REGION Network 26: Check Values
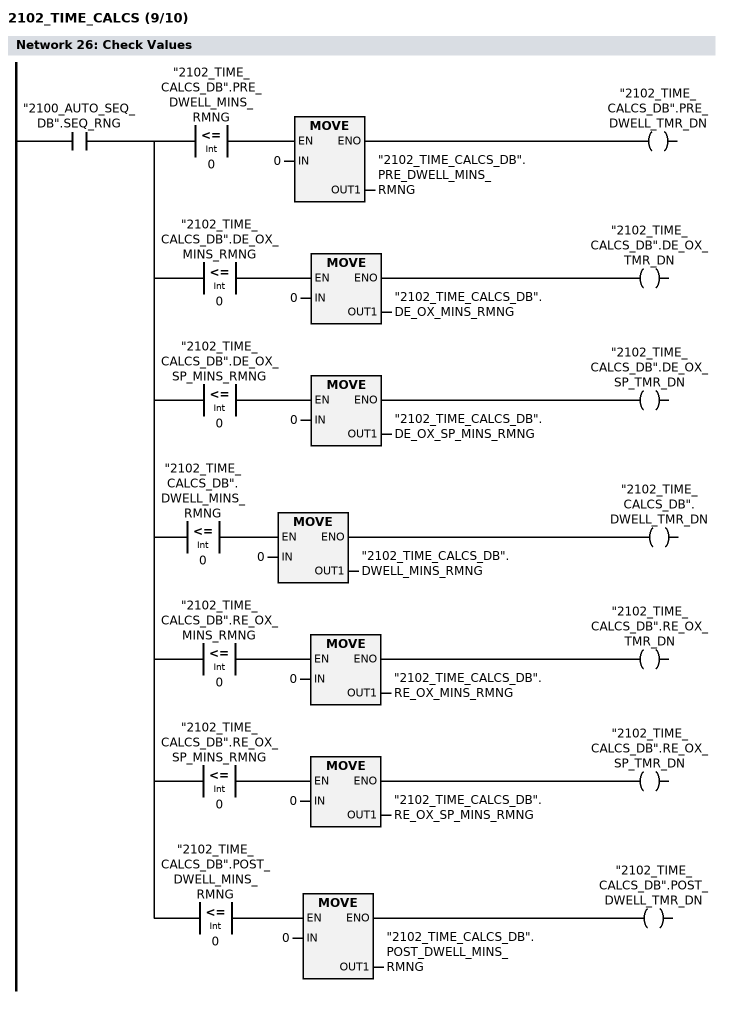
   RUNG wire#powerrail
      Contact( "2100_AUTO_SEQ_DB".SEQ_RNG )
      wire#w1
      { S7_Templates := "SrcType := Int" } LE_Contact(in1 := "2102_TIME_CALCS_DB".PRE_DWELL_MINS_RMNG, in2 := 0)
      Move(in := 0, out1 => "2102_TIME_CALCS_DB".PRE_DWELL_MINS_RMNG)
      Coil( "2102_TIME_CALCS_DB".PRE_DWELL_TMR_DN )
   END_RUNG
   RUNG wire#w1
      { S7_Templates := "SrcType := Int" } LE_Contact(in1 := "2102_TIME_CALCS_DB".DE_OX_MINS_RMNG, in2 := 0)
      Move(in := 0, out1 => "2102_TIME_CALCS_DB".DE_OX_MINS_RMNG)
      Coil( "2102_TIME_CALCS_DB".DE_OX_TMR_DN )
   END_RUNG
   RUNG wire#w1
      { S7_Templates := "SrcType := Int" } LE_Contact(in1 := "2102_TIME_CALCS_DB".DE_OX_SP_MINS_RMNG, in2 := 0)
      Move(in := 0, out1 => "2102_TIME_CALCS_DB".DE_OX_SP_MINS_RMNG)
      Coil( "2102_TIME_CALCS_DB".DE_OX_SP_TMR_DN )
   END_RUNG
   RUNG wire#w1
      { S7_Templates := "SrcType := Int" } LE_Contact(in1 := "2102_TIME_CALCS_DB".DWELL_MINS_RMNG, in2 := 0)
      Move(in := 0, out1 => "2102_TIME_CALCS_DB".DWELL_MINS_RMNG)
      Coil( "2102_TIME_CALCS_DB".DWELL_TMR_DN )
   END_RUNG
   RUNG wire#w1
      { S7_Templates := "SrcType := Int" } LE_Contact(in1 := "2102_TIME_CALCS_DB".RE_OX_MINS_RMNG, in2 := 0)
      Move(in := 0, out1 => "2102_TIME_CALCS_DB".RE_OX_MINS_RMNG)
      Coil( "2102_TIME_CALCS_DB".RE_OX_TMR_DN )
   END_RUNG
   RUNG wire#w1
      { S7_Templates := "SrcType := Int" } LE_Contact(in1 := "2102_TIME_CALCS_DB".RE_OX_SP_MINS_RMNG, in2 := 0)
      Move(in := 0, out1 => "2102_TIME_CALCS_DB".RE_OX_SP_MINS_RMNG)
      Coil( "2102_TIME_CALCS_DB".RE_OX_SP_TMR_DN )
   END_RUNG
   RUNG wire#w1
      { S7_Templates := "SrcType := Int" } LE_Contact(in1 := "2102_TIME_CALCS_DB".POST_DWELL_MINS_RMNG, in2 := 0)
      Move(in := 0, out1 => "2102_TIME_CALCS_DB".POST_DWELL_MINS_RMNG)
      Coil( "2102_TIME_CALCS_DB".POST_DWELL_TMR_DN )
   END_RUNG
   // the same network as SCL:
   #_w1 := "2100_AUTO_SEQ_DB".SEQ_RNG AND ("2102_TIME_CALCS_DB".PRE_DWELL_MINS_RMNG <= 0);
   IF #_w1 THEN "2102_TIME_CALCS_DB".PRE_DWELL_MINS_RMNG := 0; END_IF;
   "2102_TIME_CALCS_DB".PRE_DWELL_TMR_DN := #_w1;
   #_w2 := "2100_AUTO_SEQ_DB".SEQ_RNG AND ("2102_TIME_CALCS_DB".DE_OX_MINS_RMNG <= 0);
   IF #_w2 THEN "2102_TIME_CALCS_DB".DE_OX_MINS_RMNG := 0; END_IF;
   "2102_TIME_CALCS_DB".DE_OX_TMR_DN := #_w2;
   #_w3 := "2100_AUTO_SEQ_DB".SEQ_RNG AND ("2102_TIME_CALCS_DB".DE_OX_SP_MINS_RMNG <= 0);
   IF #_w3 THEN "2102_TIME_CALCS_DB".DE_OX_SP_MINS_RMNG := 0; END_IF;
   "2102_TIME_CALCS_DB".DE_OX_SP_TMR_DN := #_w3;
   #_w4 := "2100_AUTO_SEQ_DB".SEQ_RNG AND ("2102_TIME_CALCS_DB".DWELL_MINS_RMNG <= 0);
   IF #_w4 THEN "2102_TIME_CALCS_DB".DWELL_MINS_RMNG := 0; END_IF;
   "2102_TIME_CALCS_DB".DWELL_TMR_DN := #_w4;
   #_w5 := "2100_AUTO_SEQ_DB".SEQ_RNG AND ("2102_TIME_CALCS_DB".RE_OX_MINS_RMNG <= 0);
   IF #_w5 THEN "2102_TIME_CALCS_DB".RE_OX_MINS_RMNG := 0; END_IF;
   "2102_TIME_CALCS_DB".RE_OX_TMR_DN := #_w5;
   #_w6 := "2100_AUTO_SEQ_DB".SEQ_RNG AND ("2102_TIME_CALCS_DB".RE_OX_SP_MINS_RMNG <= 0);
   IF #_w6 THEN "2102_TIME_CALCS_DB".RE_OX_SP_MINS_RMNG := 0; END_IF;
   "2102_TIME_CALCS_DB".RE_OX_SP_TMR_DN := #_w6;
   #_w7 := "2100_AUTO_SEQ_DB".SEQ_RNG AND ("2102_TIME_CALCS_DB".POST_DWELL_MINS_RMNG <= 0);
   IF #_w7 THEN "2102_TIME_CALCS_DB".POST_DWELL_MINS_RMNG := 0; END_IF;
   "2102_TIME_CALCS_DB".POST_DWELL_TMR_DN := #_w7;
END_REGION

REGION Network 27: Total Remaining Time
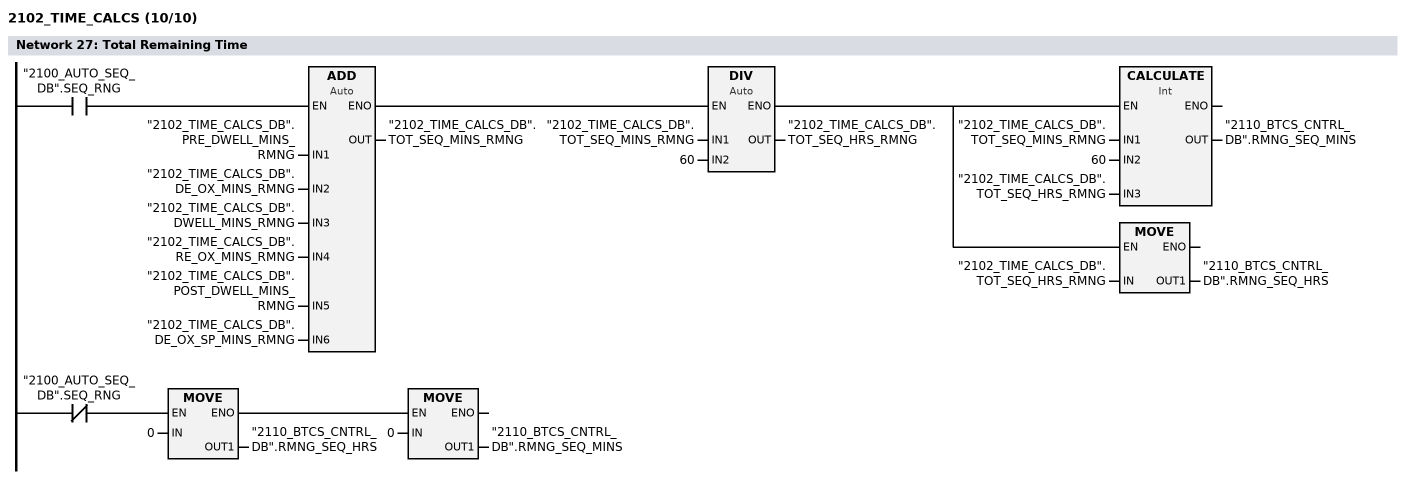
   RUNG wire#powerrail
      Contact( "2100_AUTO_SEQ_DB".SEQ_RNG )
      Add(in1 := "2102_TIME_CALCS_DB".PRE_DWELL_MINS_RMNG, in2 := "2102_TIME_CALCS_DB".DE_OX_MINS_RMNG, in3 := "2102_TIME_CALCS_DB".DWELL_MINS_RMNG, in4 := "2102_TIME_CALCS_DB".RE_OX_MINS_RMNG, in5 := "2102_TIME_CALCS_DB".POST_DWELL_MINS_RMNG, in6 := "2102_TIME_CALCS_DB".DE_OX_SP_MINS_RMNG, out => "2102_TIME_CALCS_DB".TOT_SEQ_MINS_RMNG)
      Div(in1 := "2102_TIME_CALCS_DB".TOT_SEQ_MINS_RMNG, in2 := 60, out => "2102_TIME_CALCS_DB".TOT_SEQ_HRS_RMNG)
      wire#w1
      { S7_Templates := "SrcType := Int"; S7_Expression := "IN1-(IN3*IN2)" } Calculate(in1 := "2102_TIME_CALCS_DB".TOT_SEQ_MINS_RMNG, in2 := 60, in3 := "2102_TIME_CALCS_DB".TOT_SEQ_HRS_RMNG, out => "2110_BTCS_CNTRL_DB".RMNG_SEQ_MINS)
   END_RUNG
   RUNG wire#w1
      Move(in := "2102_TIME_CALCS_DB".TOT_SEQ_HRS_RMNG, out1 => "2110_BTCS_CNTRL_DB".RMNG_SEQ_HRS)
   END_RUNG
   RUNG wire#powerrail
      I_Contact( "2100_AUTO_SEQ_DB".SEQ_RNG )
      Move(in := 0, out1 => "2110_BTCS_CNTRL_DB".RMNG_SEQ_HRS)
      Move(in := 0, out1 => "2110_BTCS_CNTRL_DB".RMNG_SEQ_MINS)
   END_RUNG
   // the same network as SCL:
   IF "2100_AUTO_SEQ_DB".SEQ_RNG THEN
       "2102_TIME_CALCS_DB".TOT_SEQ_MINS_RMNG := "2102_TIME_CALCS_DB".PRE_DWELL_MINS_RMNG + "2102_TIME_CALCS_DB".DE_OX_MINS_RMNG + "2102_TIME_CALCS_DB".DWELL_MINS_RMNG + "2102_TIME_CALCS_DB".RE_OX_MINS_RMNG + "2102_TIME_CALCS_DB".POST_DWELL_MINS_RMNG + "2102_TIME_CALCS_DB".DE_OX_SP_MINS_RMNG;
       "2102_TIME_CALCS_DB".TOT_SEQ_HRS_RMNG := "2102_TIME_CALCS_DB".TOT_SEQ_MINS_RMNG / 60;
       "2110_BTCS_CNTRL_DB".RMNG_SEQ_MINS := "2102_TIME_CALCS_DB".TOT_SEQ_MINS_RMNG-("2102_TIME_CALCS_DB".TOT_SEQ_HRS_RMNG*60);
       "2110_BTCS_CNTRL_DB".RMNG_SEQ_HRS := "2102_TIME_CALCS_DB".TOT_SEQ_HRS_RMNG;
   END_IF;
   IF NOT "2100_AUTO_SEQ_DB".SEQ_RNG THEN
       "2110_BTCS_CNTRL_DB".RMNG_SEQ_HRS := 0;
       "2110_BTCS_CNTRL_DB".RMNG_SEQ_MINS := 0;
   END_IF;
END_REGION
END_FUNCTION

FUNCTION "2110_BTCS_CNTRL" : Void   // FC2110, LAD
TITLE = Barge Tank Control System
{ S7_Optimized_Access := 'TRUE' }
AUTHOR : JRS
VERSION : 0.1
// For running the optional barge tank control system
BEGIN

REGION Network 1: Automatic Commands
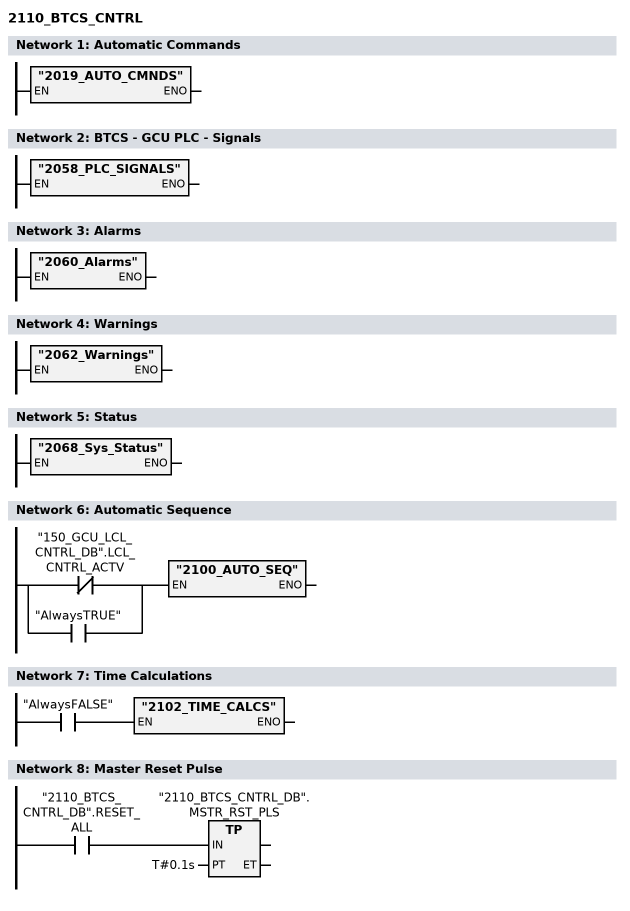
   RUNG wire#powerrail
      "2019_AUTO_CMNDS"()
   END_RUNG
   // the same network as SCL:
   "2019_AUTO_CMNDS"();
END_REGION

REGION Network 2: BTCS - GCU PLC - Signals
   RUNG wire#powerrail
      "2058_PLC_SIGNALS"()
   END_RUNG
   // the same network as SCL:
   "2058_PLC_SIGNALS"();
END_REGION

REGION Network 3: Alarms
   RUNG wire#powerrail
      "2060_Alarms"()
   END_RUNG
   // the same network as SCL:
   "2060_Alarms"();
END_REGION

REGION Network 4: Warnings
   RUNG wire#powerrail
      "2062_Warnings"()
   END_RUNG
   // the same network as SCL:
   "2062_Warnings"();
END_REGION

REGION Network 5: Status
   RUNG wire#powerrail
      "2068_Sys_Status"()
   END_RUNG
   // the same network as SCL:
   "2068_Sys_Status"();
END_REGION

REGION Network 6: Automatic Sequence
   RUNG wire#powerrail
      I_Contact( "150_GCU_LCL_CNTRL_DB".LCL_CNTRL_ACTV )
      wire#w1
      "2100_AUTO_SEQ"()
   END_RUNG
   RUNG wire#powerrail
      Contact( "AlwaysTRUE" )
   END_RUNG wire#w1
   // the same network as SCL:
   IF NOT "150_GCU_LCL_CNTRL_DB".LCL_CNTRL_ACTV OR "AlwaysTRUE" THEN "2100_AUTO_SEQ"(); END_IF;
END_REGION

REGION Network 7: Time Calculations
   RUNG wire#powerrail
      Contact( "AlwaysFALSE" )
      "2102_TIME_CALCS"()
   END_RUNG
   // the same network as SCL:
   IF "AlwaysFALSE" THEN "2102_TIME_CALCS"(); END_IF;
END_REGION

REGION Network 8: Master Reset Pulse
   "2110_BTCS_CNTRL_DB".MSTR_RST_PLS.TP(IN := "2110_BTCS_CNTRL_DB".RESET_ALL, PT := T#0.1s);
END_REGION
END_FUNCTION

// folder: 300 - 499 Counter and Timer DBs

FUNCTION "300_AUT_SEQ_TIMERS" : Void   // FC300, LAD
TITLE = Automatic Sequence Timers
{ S7_Optimized_Access := 'TRUE' }
AUTHOR : JRS
VERSION : 0.1
// For specific sequence timers not covered by step FB timers
BEGIN

REGION Network 1: Pre GCU Start Command Delay (CV341 Closed)
   // Get time value from HMI data
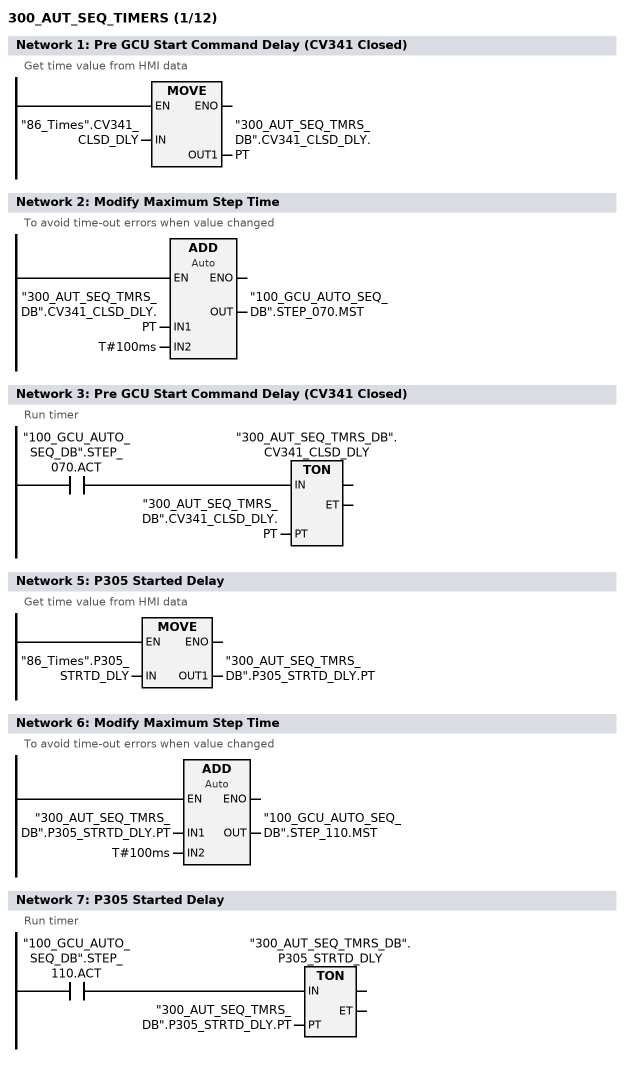
   RUNG wire#powerrail
      Move(in := "86_Times".CV341_CLSD_DLY, out1 => "300_AUT_SEQ_TMRS_DB".CV341_CLSD_DLY.PT)
   END_RUNG
   // the same network as SCL:
   "300_AUT_SEQ_TMRS_DB".CV341_CLSD_DLY.PT := "86_Times".CV341_CLSD_DLY;
END_REGION

REGION Network 2: Modify Maximum Step Time
   // To avoid time-out errors when value changed
   RUNG wire#powerrail
      Add(in1 := "300_AUT_SEQ_TMRS_DB".CV341_CLSD_DLY.PT, in2 := T#100ms, out => "100_GCU_AUTO_SEQ_DB".STEP_070.MST)
   END_RUNG
   // the same network as SCL:
   "100_GCU_AUTO_SEQ_DB".STEP_070.MST := "300_AUT_SEQ_TMRS_DB".CV341_CLSD_DLY.PT + T#100ms;
END_REGION

REGION Network 3: Pre GCU Start Command Delay (CV341 Closed)
   // Run timer
   "300_AUT_SEQ_TMRS_DB".CV341_CLSD_DLY.TON(IN := "100_GCU_AUTO_SEQ_DB".STEP_070.ACT,
                           PT := "300_AUT_SEQ_TMRS_DB".CV341_CLSD_DLY.PT);
END_REGION

REGION Network 5: P305 Started Delay
   // Get time value from HMI data
   RUNG wire#powerrail
      Move(in := "86_Times".P305_STRTD_DLY, out1 => "300_AUT_SEQ_TMRS_DB".P305_STRTD_DLY.PT)
   END_RUNG
   // the same network as SCL:
   "300_AUT_SEQ_TMRS_DB".P305_STRTD_DLY.PT := "86_Times".P305_STRTD_DLY;
END_REGION

REGION Network 6: Modify Maximum Step Time
   // To avoid time-out errors when value changed
   RUNG wire#powerrail
      Add(in1 := "300_AUT_SEQ_TMRS_DB".P305_STRTD_DLY.PT, in2 := T#100ms, out => "100_GCU_AUTO_SEQ_DB".STEP_110.MST)
   END_RUNG
   // the same network as SCL:
   "100_GCU_AUTO_SEQ_DB".STEP_110.MST := "300_AUT_SEQ_TMRS_DB".P305_STRTD_DLY.PT + T#100ms;
END_REGION

REGION Network 7: P305 Started Delay
   // Run timer
   "300_AUT_SEQ_TMRS_DB".P305_STRTD_DLY.TON(IN := "100_GCU_AUTO_SEQ_DB".STEP_110.ACT,
                           PT := "300_AUT_SEQ_TMRS_DB".P305_STRTD_DLY.PT);
END_REGION

REGION Network 9: P304 Started Delay
   // Get time value from HMI data
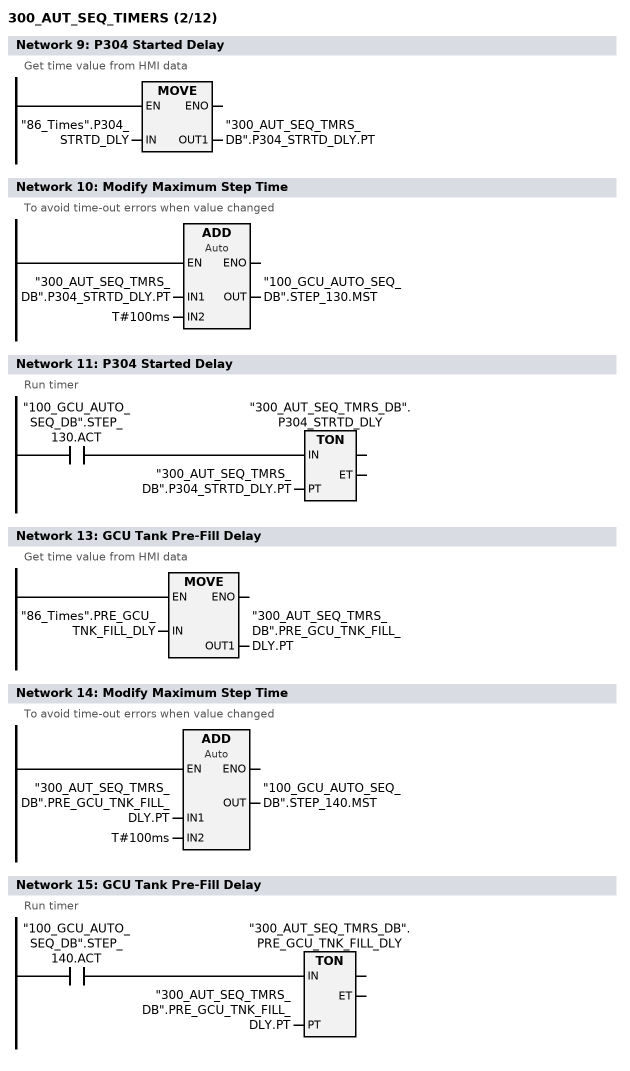
   RUNG wire#powerrail
      Move(in := "86_Times".P304_STRTD_DLY, out1 => "300_AUT_SEQ_TMRS_DB".P304_STRTD_DLY.PT)
   END_RUNG
   // the same network as SCL:
   "300_AUT_SEQ_TMRS_DB".P304_STRTD_DLY.PT := "86_Times".P304_STRTD_DLY;
END_REGION

REGION Network 10: Modify Maximum Step Time
   // To avoid time-out errors when value changed
   RUNG wire#powerrail
      Add(in1 := "300_AUT_SEQ_TMRS_DB".P304_STRTD_DLY.PT, in2 := T#100ms, out => "100_GCU_AUTO_SEQ_DB".STEP_130.MST)
   END_RUNG
   // the same network as SCL:
   "100_GCU_AUTO_SEQ_DB".STEP_130.MST := "300_AUT_SEQ_TMRS_DB".P304_STRTD_DLY.PT + T#100ms;
END_REGION

REGION Network 11: P304 Started Delay
   // Run timer
   "300_AUT_SEQ_TMRS_DB".P304_STRTD_DLY.TON(IN := "100_GCU_AUTO_SEQ_DB".STEP_130.ACT,
                           PT := "300_AUT_SEQ_TMRS_DB".P304_STRTD_DLY.PT);
END_REGION

REGION Network 13: GCU Tank Pre-Fill Delay
   // Get time value from HMI data
   RUNG wire#powerrail
      Move(in := "86_Times".PRE_GCU_TNK_FILL_DLY, out1 => "300_AUT_SEQ_TMRS_DB".PRE_GCU_TNK_FILL_DLY.PT)
   END_RUNG
   // the same network as SCL:
   "300_AUT_SEQ_TMRS_DB".PRE_GCU_TNK_FILL_DLY.PT := "86_Times".PRE_GCU_TNK_FILL_DLY;
END_REGION

REGION Network 14: Modify Maximum Step Time
   // To avoid time-out errors when value changed
   RUNG wire#powerrail
      Add(in1 := "300_AUT_SEQ_TMRS_DB".PRE_GCU_TNK_FILL_DLY.PT, in2 := T#100ms, out => "100_GCU_AUTO_SEQ_DB".STEP_140.MST)
   END_RUNG
   // the same network as SCL:
   "100_GCU_AUTO_SEQ_DB".STEP_140.MST := "300_AUT_SEQ_TMRS_DB".PRE_GCU_TNK_FILL_DLY.PT + T#100ms;
END_REGION

REGION Network 15: GCU Tank Pre-Fill Delay
   // Run timer
   "300_AUT_SEQ_TMRS_DB".PRE_GCU_TNK_FILL_DLY.TON(IN := "100_GCU_AUTO_SEQ_DB".STEP_140.ACT,
                           PT := "300_AUT_SEQ_TMRS_DB".PRE_GCU_TNK_FILL_DLY.PT);
END_REGION

REGION Network 17: GCU Tank Max Fill Time
   // Get time value from HMI data
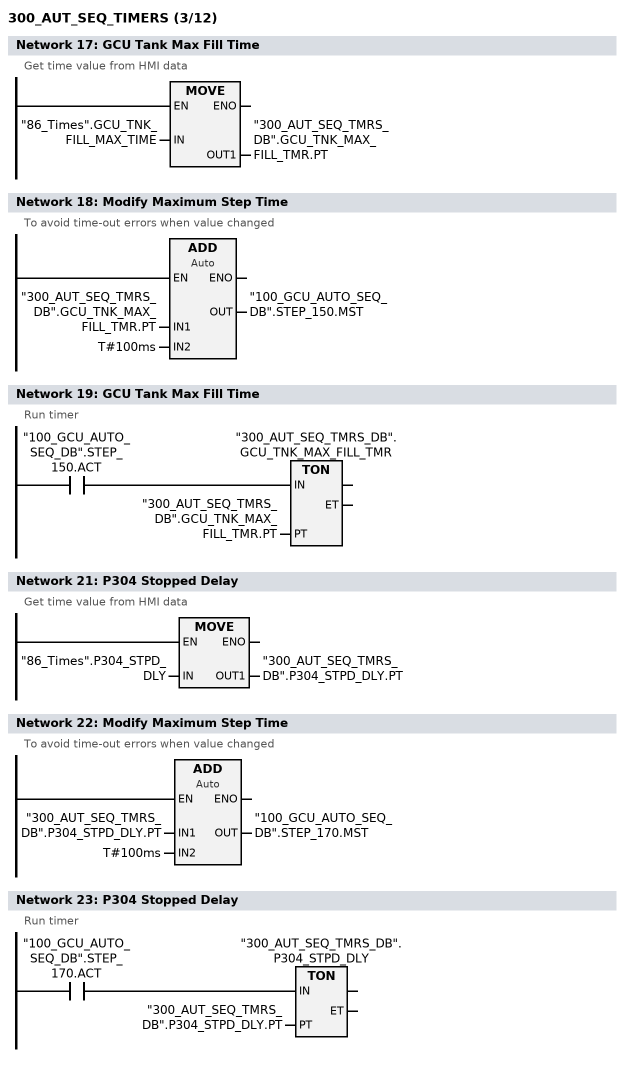
   RUNG wire#powerrail
      Move(in := "86_Times".GCU_TNK_FILL_MAX_TIME, out1 => "300_AUT_SEQ_TMRS_DB".GCU_TNK_MAX_FILL_TMR.PT)
   END_RUNG
   // the same network as SCL:
   "300_AUT_SEQ_TMRS_DB".GCU_TNK_MAX_FILL_TMR.PT := "86_Times".GCU_TNK_FILL_MAX_TIME;
END_REGION

REGION Network 18: Modify Maximum Step Time
   // To avoid time-out errors when value changed
   RUNG wire#powerrail
      Add(in1 := "300_AUT_SEQ_TMRS_DB".GCU_TNK_MAX_FILL_TMR.PT, in2 := T#100ms, out => "100_GCU_AUTO_SEQ_DB".STEP_150.MST)
   END_RUNG
   // the same network as SCL:
   "100_GCU_AUTO_SEQ_DB".STEP_150.MST := "300_AUT_SEQ_TMRS_DB".GCU_TNK_MAX_FILL_TMR.PT + T#100ms;
END_REGION

REGION Network 19: GCU Tank Max Fill Time
   // Run timer
   "300_AUT_SEQ_TMRS_DB".GCU_TNK_MAX_FILL_TMR.TON(IN := "100_GCU_AUTO_SEQ_DB".STEP_150.ACT,
                           PT := "300_AUT_SEQ_TMRS_DB".GCU_TNK_MAX_FILL_TMR.PT);
END_REGION

REGION Network 21: P304 Stopped Delay
   // Get time value from HMI data
   RUNG wire#powerrail
      Move(in := "86_Times".P304_STPD_DLY, out1 => "300_AUT_SEQ_TMRS_DB".P304_STPD_DLY.PT)
   END_RUNG
   // the same network as SCL:
   "300_AUT_SEQ_TMRS_DB".P304_STPD_DLY.PT := "86_Times".P304_STPD_DLY;
END_REGION

REGION Network 22: Modify Maximum Step Time
   // To avoid time-out errors when value changed
   RUNG wire#powerrail
      Add(in1 := "300_AUT_SEQ_TMRS_DB".P304_STPD_DLY.PT, in2 := T#100ms, out => "100_GCU_AUTO_SEQ_DB".STEP_170.MST)
   END_RUNG
   // the same network as SCL:
   "100_GCU_AUTO_SEQ_DB".STEP_170.MST := "300_AUT_SEQ_TMRS_DB".P304_STPD_DLY.PT + T#100ms;
END_REGION

REGION Network 23: P304 Stopped Delay
   // Run timer
   "300_AUT_SEQ_TMRS_DB".P304_STPD_DLY.TON(IN := "100_GCU_AUTO_SEQ_DB".STEP_170.ACT,
                           PT := "300_AUT_SEQ_TMRS_DB".P304_STPD_DLY.PT);
END_REGION

REGION Network 25: P305 Stopped Delay
   // Get time value from HMI data
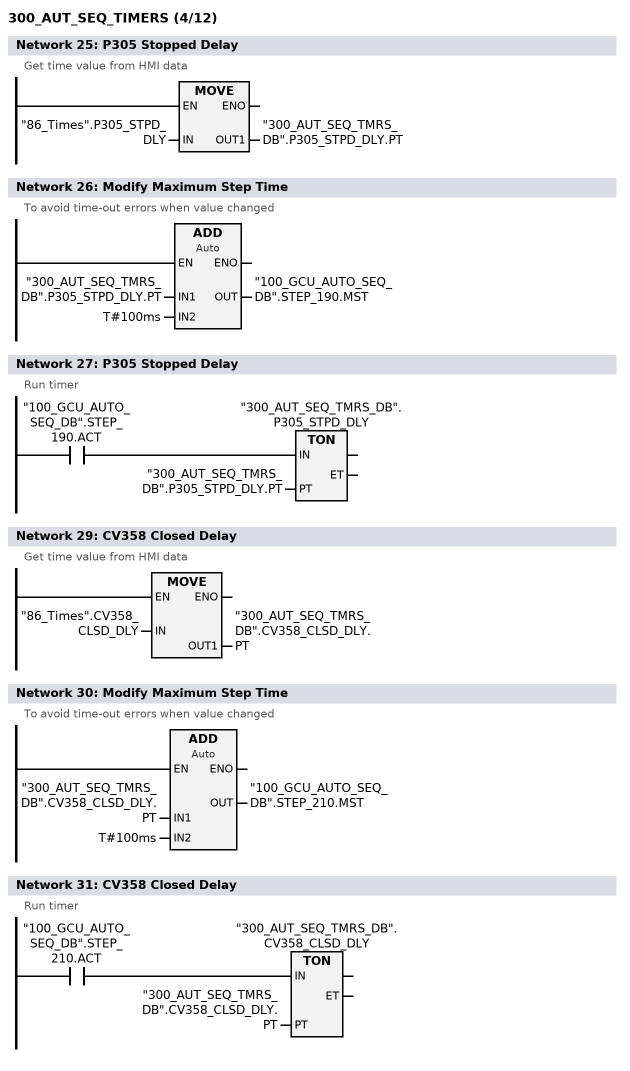
   RUNG wire#powerrail
      Move(in := "86_Times".P305_STPD_DLY, out1 => "300_AUT_SEQ_TMRS_DB".P305_STPD_DLY.PT)
   END_RUNG
   // the same network as SCL:
   "300_AUT_SEQ_TMRS_DB".P305_STPD_DLY.PT := "86_Times".P305_STPD_DLY;
END_REGION

REGION Network 26: Modify Maximum Step Time
   // To avoid time-out errors when value changed
   RUNG wire#powerrail
      Add(in1 := "300_AUT_SEQ_TMRS_DB".P305_STPD_DLY.PT, in2 := T#100ms, out => "100_GCU_AUTO_SEQ_DB".STEP_190.MST)
   END_RUNG
   // the same network as SCL:
   "100_GCU_AUTO_SEQ_DB".STEP_190.MST := "300_AUT_SEQ_TMRS_DB".P305_STPD_DLY.PT + T#100ms;
END_REGION

REGION Network 27: P305 Stopped Delay
   // Run timer
   "300_AUT_SEQ_TMRS_DB".P305_STPD_DLY.TON(IN := "100_GCU_AUTO_SEQ_DB".STEP_190.ACT,
                           PT := "300_AUT_SEQ_TMRS_DB".P305_STPD_DLY.PT);
END_REGION

REGION Network 29: CV358 Closed Delay
   // Get time value from HMI data
   RUNG wire#powerrail
      Move(in := "86_Times".CV358_CLSD_DLY, out1 => "300_AUT_SEQ_TMRS_DB".CV358_CLSD_DLY.PT)
   END_RUNG
   // the same network as SCL:
   "300_AUT_SEQ_TMRS_DB".CV358_CLSD_DLY.PT := "86_Times".CV358_CLSD_DLY;
END_REGION

REGION Network 30: Modify Maximum Step Time
   // To avoid time-out errors when value changed
   RUNG wire#powerrail
      Add(in1 := "300_AUT_SEQ_TMRS_DB".CV358_CLSD_DLY.PT, in2 := T#100ms, out => "100_GCU_AUTO_SEQ_DB".STEP_210.MST)
   END_RUNG
   // the same network as SCL:
   "100_GCU_AUTO_SEQ_DB".STEP_210.MST := "300_AUT_SEQ_TMRS_DB".CV358_CLSD_DLY.PT + T#100ms;
END_REGION

REGION Network 31: CV358 Closed Delay
   // Run timer
   "300_AUT_SEQ_TMRS_DB".CV358_CLSD_DLY.TON(IN := "100_GCU_AUTO_SEQ_DB".STEP_210.ACT,
                           PT := "300_AUT_SEQ_TMRS_DB".CV358_CLSD_DLY.PT);
END_REGION

REGION Network 33: P303 Started Delay
   // Get time value from HMI data
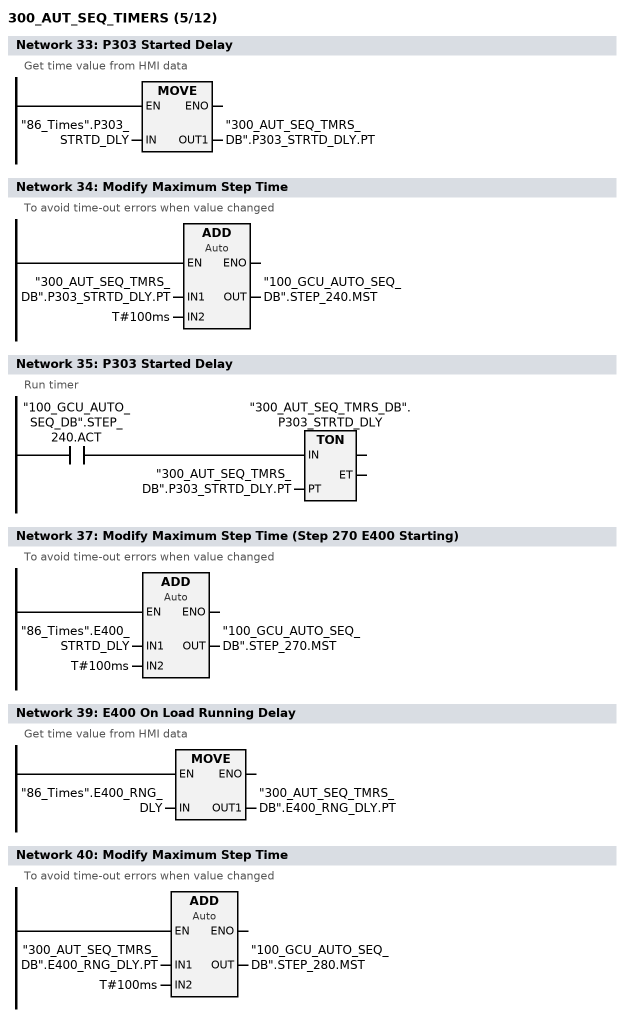
   RUNG wire#powerrail
      Move(in := "86_Times".P303_STRTD_DLY, out1 => "300_AUT_SEQ_TMRS_DB".P303_STRTD_DLY.PT)
   END_RUNG
   // the same network as SCL:
   "300_AUT_SEQ_TMRS_DB".P303_STRTD_DLY.PT := "86_Times".P303_STRTD_DLY;
END_REGION

REGION Network 34: Modify Maximum Step Time
   // To avoid time-out errors when value changed
   RUNG wire#powerrail
      Add(in1 := "300_AUT_SEQ_TMRS_DB".P303_STRTD_DLY.PT, in2 := T#100ms, out => "100_GCU_AUTO_SEQ_DB".STEP_240.MST)
   END_RUNG
   // the same network as SCL:
   "100_GCU_AUTO_SEQ_DB".STEP_240.MST := "300_AUT_SEQ_TMRS_DB".P303_STRTD_DLY.PT + T#100ms;
END_REGION

REGION Network 35: P303 Started Delay
   // Run timer
   "300_AUT_SEQ_TMRS_DB".P303_STRTD_DLY.TON(IN := "100_GCU_AUTO_SEQ_DB".STEP_240.ACT,
                           PT := "300_AUT_SEQ_TMRS_DB".P303_STRTD_DLY.PT);
END_REGION

REGION Network 37: Modify Maximum Step Time (Step 270 E400 Starting)
   // To avoid time-out errors when value changed
   RUNG wire#powerrail
      Add(in1 := "86_Times".E400_STRTD_DLY, in2 := T#100ms, out => "100_GCU_AUTO_SEQ_DB".STEP_270.MST)
   END_RUNG
   // the same network as SCL:
   "100_GCU_AUTO_SEQ_DB".STEP_270.MST := "86_Times".E400_STRTD_DLY + T#100ms;
END_REGION

REGION Network 39: E400 On Load Running Delay
   // Get time value from HMI data
   RUNG wire#powerrail
      Move(in := "86_Times".E400_RNG_DLY, out1 => "300_AUT_SEQ_TMRS_DB".E400_RNG_DLY.PT)
   END_RUNG
   // the same network as SCL:
   "300_AUT_SEQ_TMRS_DB".E400_RNG_DLY.PT := "86_Times".E400_RNG_DLY;
END_REGION

REGION Network 40: Modify Maximum Step Time
   // To avoid time-out errors when value changed
   RUNG wire#powerrail
      Add(in1 := "300_AUT_SEQ_TMRS_DB".E400_RNG_DLY.PT, in2 := T#100ms, out => "100_GCU_AUTO_SEQ_DB".STEP_280.MST)
   END_RUNG
   // the same network as SCL:
   "100_GCU_AUTO_SEQ_DB".STEP_280.MST := "300_AUT_SEQ_TMRS_DB".E400_RNG_DLY.PT + T#100ms;
END_REGION

REGION Network 41: E400 On Load Running Delay
   // Run timer
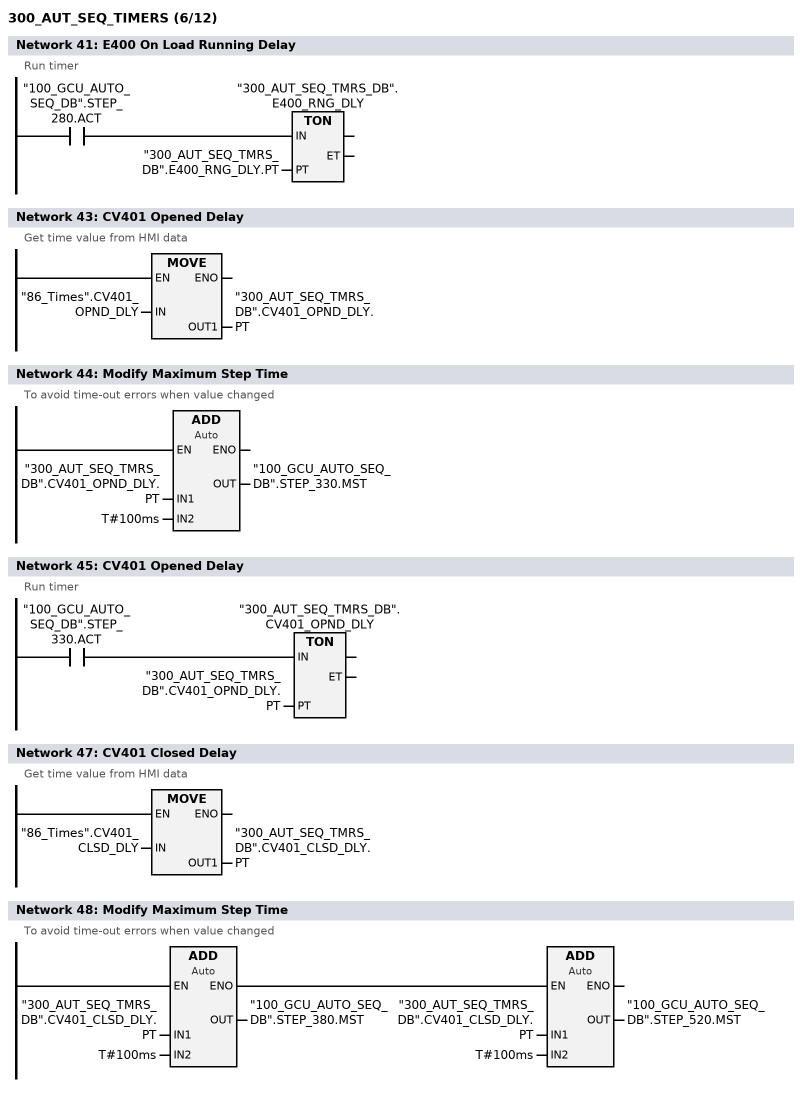
   "300_AUT_SEQ_TMRS_DB".E400_RNG_DLY.TON(IN := "100_GCU_AUTO_SEQ_DB".STEP_280.ACT,
                           PT := "300_AUT_SEQ_TMRS_DB".E400_RNG_DLY.PT);
END_REGION

REGION Network 43: CV401 Opened Delay
   // Get time value from HMI data
   RUNG wire#powerrail
      Move(in := "86_Times".CV401_OPND_DLY, out1 => "300_AUT_SEQ_TMRS_DB".CV401_OPND_DLY.PT)
   END_RUNG
   // the same network as SCL:
   "300_AUT_SEQ_TMRS_DB".CV401_OPND_DLY.PT := "86_Times".CV401_OPND_DLY;
END_REGION

REGION Network 44: Modify Maximum Step Time
   // To avoid time-out errors when value changed
   RUNG wire#powerrail
      Add(in1 := "300_AUT_SEQ_TMRS_DB".CV401_OPND_DLY.PT, in2 := T#100ms, out => "100_GCU_AUTO_SEQ_DB".STEP_330.MST)
   END_RUNG
   // the same network as SCL:
   "100_GCU_AUTO_SEQ_DB".STEP_330.MST := "300_AUT_SEQ_TMRS_DB".CV401_OPND_DLY.PT + T#100ms;
END_REGION

REGION Network 45: CV401 Opened Delay
   // Run timer
   "300_AUT_SEQ_TMRS_DB".CV401_OPND_DLY.TON(IN := "100_GCU_AUTO_SEQ_DB".STEP_330.ACT,
                           PT := "300_AUT_SEQ_TMRS_DB".CV401_OPND_DLY.PT);
END_REGION

REGION Network 47: CV401 Closed Delay
   // Get time value from HMI data
   RUNG wire#powerrail
      Move(in := "86_Times".CV401_CLSD_DLY, out1 => "300_AUT_SEQ_TMRS_DB".CV401_CLSD_DLY.PT)
   END_RUNG
   // the same network as SCL:
   "300_AUT_SEQ_TMRS_DB".CV401_CLSD_DLY.PT := "86_Times".CV401_CLSD_DLY;
END_REGION

REGION Network 48: Modify Maximum Step Time
   // To avoid time-out errors when value changed
   RUNG wire#powerrail
      Add(in1 := "300_AUT_SEQ_TMRS_DB".CV401_CLSD_DLY.PT, in2 := T#100ms, out => "100_GCU_AUTO_SEQ_DB".STEP_380.MST)
      Add(in1 := "300_AUT_SEQ_TMRS_DB".CV401_CLSD_DLY.PT, in2 := T#100ms, out => "100_GCU_AUTO_SEQ_DB".STEP_520.MST)
   END_RUNG
   // the same network as SCL:
   "100_GCU_AUTO_SEQ_DB".STEP_380.MST := "300_AUT_SEQ_TMRS_DB".CV401_CLSD_DLY.PT + T#100ms;
   "100_GCU_AUTO_SEQ_DB".STEP_520.MST := "300_AUT_SEQ_TMRS_DB".CV401_CLSD_DLY.PT + T#100ms;
END_REGION

REGION Network 49: CV401 Closed Delay
   // Run timer
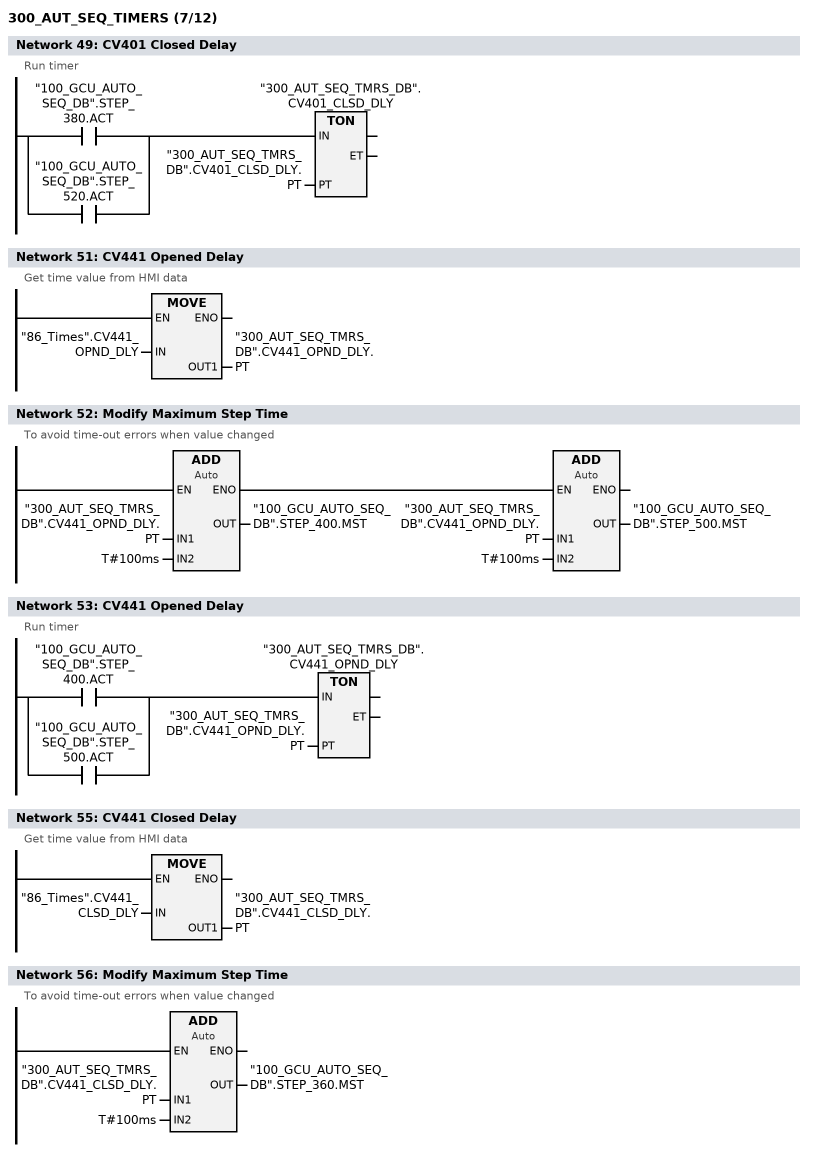
   "300_AUT_SEQ_TMRS_DB".CV401_CLSD_DLY.TON(IN := "100_GCU_AUTO_SEQ_DB".STEP_380.ACT OR "100_GCU_AUTO_SEQ_DB".STEP_520.ACT,
                           PT := "300_AUT_SEQ_TMRS_DB".CV401_CLSD_DLY.PT);
END_REGION

REGION Network 51: CV441 Opened Delay
   // Get time value from HMI data
   RUNG wire#powerrail
      Move(in := "86_Times".CV441_OPND_DLY, out1 => "300_AUT_SEQ_TMRS_DB".CV441_OPND_DLY.PT)
   END_RUNG
   // the same network as SCL:
   "300_AUT_SEQ_TMRS_DB".CV441_OPND_DLY.PT := "86_Times".CV441_OPND_DLY;
END_REGION

REGION Network 52: Modify Maximum Step Time
   // To avoid time-out errors when value changed
   RUNG wire#powerrail
      Add(in1 := "300_AUT_SEQ_TMRS_DB".CV441_OPND_DLY.PT, in2 := T#100ms, out => "100_GCU_AUTO_SEQ_DB".STEP_400.MST)
      Add(in1 := "300_AUT_SEQ_TMRS_DB".CV441_OPND_DLY.PT, in2 := T#100ms, out => "100_GCU_AUTO_SEQ_DB".STEP_500.MST)
   END_RUNG
   // the same network as SCL:
   "100_GCU_AUTO_SEQ_DB".STEP_400.MST := "300_AUT_SEQ_TMRS_DB".CV441_OPND_DLY.PT + T#100ms;
   "100_GCU_AUTO_SEQ_DB".STEP_500.MST := "300_AUT_SEQ_TMRS_DB".CV441_OPND_DLY.PT + T#100ms;
END_REGION

REGION Network 53: CV441 Opened Delay
   // Run timer
   "300_AUT_SEQ_TMRS_DB".CV441_OPND_DLY.TON(IN := "100_GCU_AUTO_SEQ_DB".STEP_400.ACT OR "100_GCU_AUTO_SEQ_DB".STEP_500.ACT,
                           PT := "300_AUT_SEQ_TMRS_DB".CV441_OPND_DLY.PT);
END_REGION

REGION Network 55: CV441 Closed Delay
   // Get time value from HMI data
   RUNG wire#powerrail
      Move(in := "86_Times".CV441_CLSD_DLY, out1 => "300_AUT_SEQ_TMRS_DB".CV441_CLSD_DLY.PT)
   END_RUNG
   // the same network as SCL:
   "300_AUT_SEQ_TMRS_DB".CV441_CLSD_DLY.PT := "86_Times".CV441_CLSD_DLY;
END_REGION

REGION Network 56: Modify Maximum Step Time
   // To avoid time-out errors when value changed
   RUNG wire#powerrail
      Add(in1 := "300_AUT_SEQ_TMRS_DB".CV441_CLSD_DLY.PT, in2 := T#100ms, out => "100_GCU_AUTO_SEQ_DB".STEP_360.MST)
   END_RUNG
   // the same network as SCL:
   "100_GCU_AUTO_SEQ_DB".STEP_360.MST := "300_AUT_SEQ_TMRS_DB".CV441_CLSD_DLY.PT + T#100ms;
END_REGION

REGION Network 57: CV441 Closed Delay
   // Run timer
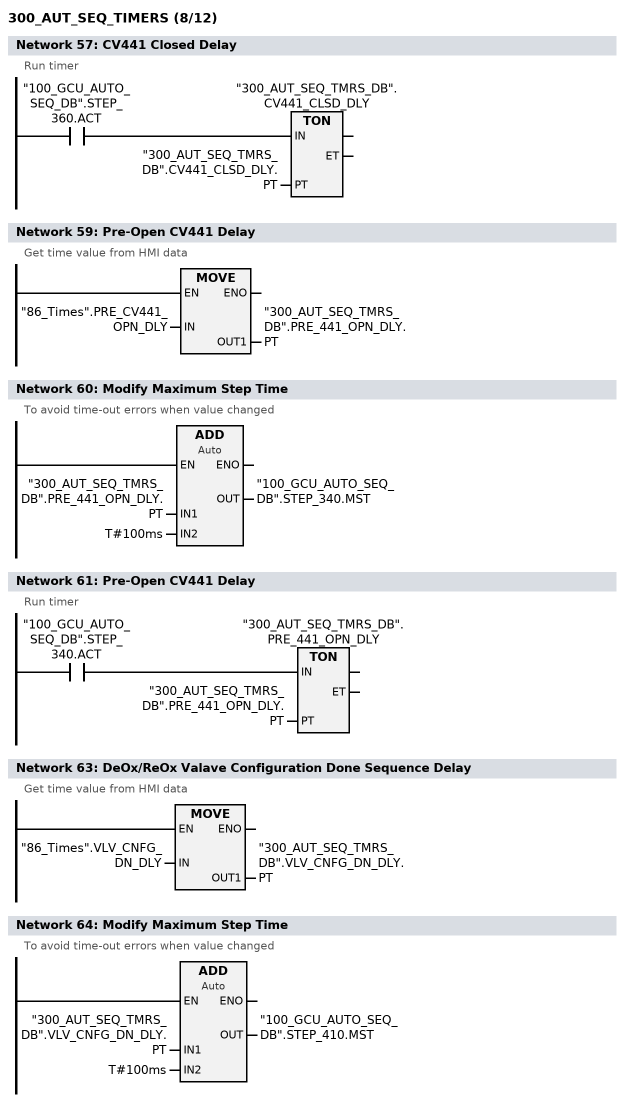
   "300_AUT_SEQ_TMRS_DB".CV441_CLSD_DLY.TON(IN := "100_GCU_AUTO_SEQ_DB".STEP_360.ACT,
                           PT := "300_AUT_SEQ_TMRS_DB".CV441_CLSD_DLY.PT);
END_REGION

REGION Network 59: Pre-Open CV441 Delay
   // Get time value from HMI data
   RUNG wire#powerrail
      Move(in := "86_Times".PRE_CV441_OPN_DLY, out1 => "300_AUT_SEQ_TMRS_DB".PRE_441_OPN_DLY.PT)
   END_RUNG
   // the same network as SCL:
   "300_AUT_SEQ_TMRS_DB".PRE_441_OPN_DLY.PT := "86_Times".PRE_CV441_OPN_DLY;
END_REGION

REGION Network 60: Modify Maximum Step Time
   // To avoid time-out errors when value changed
   RUNG wire#powerrail
      Add(in1 := "300_AUT_SEQ_TMRS_DB".PRE_441_OPN_DLY.PT, in2 := T#100ms, out => "100_GCU_AUTO_SEQ_DB".STEP_340.MST)
   END_RUNG
   // the same network as SCL:
   "100_GCU_AUTO_SEQ_DB".STEP_340.MST := "300_AUT_SEQ_TMRS_DB".PRE_441_OPN_DLY.PT + T#100ms;
END_REGION

REGION Network 61: Pre-Open CV441 Delay
   // Run timer
   "300_AUT_SEQ_TMRS_DB".PRE_441_OPN_DLY.TON(IN := "100_GCU_AUTO_SEQ_DB".STEP_340.ACT,
                           PT := "300_AUT_SEQ_TMRS_DB".PRE_441_OPN_DLY.PT);
END_REGION
